   4491: 'Carrier 70 Standard Input Card Fault', class No Acknowledgement, trigger "DB302_HMI_Faults_Carrier70_Faults_0" bit 10
   4492: 'Carrier 70 Standard Output Card Fault', class No Acknowledgement, trigger "DB302_HMI_Faults_Carrier70_Faults_0" bit 11
   4493: 'Carrier 70 Encoder Position Fault', class No Acknowledgement, trigger "DB302_HMI_Faults_Carrier70_Faults_0" bit 12
   4494: 'Carrier 70 Encoder Internal Error', class No Acknowledgement, trigger "DB302_HMI_Faults_Carrier70_Faults_0" bit 13
   4495: 'Carrier 70 Encoder Comm Fault', class No Acknowledgement, trigger "DB302_HMI_Faults_Carrier70_Faults_0" bit 14
   4496: 'Carrier 70 HMI Comm Fault', class No Acknowledgement, trigger "DB302_HMI_Faults_Carrier70_Faults_0" bit 15
   4497: 'Carrier 70 Crash Detection Fault', class No Acknowledgement, trigger "DB302_HMI_Faults_Carrier70_Faults_1" bit 0
   4498: 'Carrier 70 Carrier Number Invalid', class No Acknowledgement, trigger "DB302_HMI_Faults_Carrier70_Faults_1" bit 1
   4499: 'Carrier 70 Drive: PROFINET configuration error', class No Acknowledgement, trigger "DB302_HMI_Faults_Carrier70_Faults_1" bit 2
   4500: 'Carrier 70 Drive: Error internal communications', class No Acknowledgement, trigger "DB302_HMI_Faults_Carrier70_Faults_1" bit 3
   4501: 'Carrier 70 Drive: Motor overtemperature', class No Acknowledgement, trigger "DB302_HMI_Faults_Carrier70_Faults_1" bit 4
   4502: 'Carrier 70 Drive: Motor overcurrent', class No Acknowledgement, trigger "DB302_HMI_Faults_Carrier70_Faults_1" bit 5
   4503: 'Carrier 70 Drive: Infeed or power unit not ready', class No Acknowledgement, trigger "DB302_HMI_Faults_Carrier70_Faults_1" bit 6
   4504: 'Carrier 70 Drive: Short-circuit/ground fault detected', class No Acknowledgement, trigger "DB302_HMI_Faults_Carrier70_Faults_1" bit 7
   4505: 'Carrier 70 Drive: PROFINET Setpoint timeout', class No Acknowledgement, trigger "DB302_HMI_Faults_Carrier70_Faults_1" bit 8
   4506: 'Carrier 70 Power unit: Overcurrent', class No Acknowledgement, trigger "DB302_HMI_Faults_Carrier70_Faults_1" bit 9
   4507: 'Carrier 70 Power unit: DC link voltage overvoltage', class No Acknowledgement, trigger "DB302_HMI_Faults_Carrier70_Faults_1" bit 10
   4508: 'Carrier 70 Power unit: DC link voltage undervoltage', class No Acknowledgement, trigger "DB302_HMI_Faults_Carrier70_Faults_1" bit 11
   4509: 'Carrier 70 Power unit: Line phase failure in main circuit', class No Acknowledgement, trigger "DB302_HMI_Faults_Carrier70_Faults_1" bit 12
   4510: 'Carrier 70 Power unit: Phase failure motor cable', class No Acknowledgement, trigger "DB302_HMI_Faults_Carrier70_Faults_1" bit 13
   4511: 'Carrier 70 Power unit: Ground fault', class No Acknowledgement, trigger "DB302_HMI_Faults_Carrier70_Faults_1" bit 14
   4512: 'Spare_Fault_4512', class No Acknowledgement, trigger "DB302_HMI_Faults_Carrier70_Faults_1" bit 15
   4513: 'Carrier 70 Motion Off Fault', class No Acknowledgement, trigger "DB302_HMI_Faults_Carrier70_Faults_2" bit 0
   4514: 'Carrier 70 Motion On Fault', class No Acknowledgement, trigger "DB302_HMI_Faults_Carrier70_Faults_2" bit 1
   4515: 'Carrier 70 Spacing Fault', class No Acknowledgement, trigger "DB302_HMI_Faults_Carrier70_Faults_2" bit 2
   4516: 'Carrier 70 Duplicate Carrier Number Fault', class No Acknowledgement, trigger "DB302_HMI_Faults_Carrier70_Faults_2" bit 3
   4517: 'Spare_Fault_4517', class No Acknowledgement, trigger "DB302_HMI_Faults_Carrier70_Faults_2" bit 4
   4518: 'Spare_Fault_4518', class No Acknowledgement, trigger "DB302_HMI_Faults_Carrier70_Faults_2" bit 5
   4519: 'Spare_Fault_4519', class No Acknowledgement, trigger "DB302_HMI_Faults_Carrier70_Faults_2" bit 6
   4520: 'Spare_Fault_4520', class No Acknowledgement, trigger "DB302_HMI_Faults_Carrier70_Faults_2" bit 7
   4521: 'Spare_Fault_4521', class No Acknowledgement, trigger "DB302_HMI_Faults_Carrier70_Faults_2" bit 8
   4522: 'Spare_Fault_4522', class No Acknowledgement, trigger "DB302_HMI_Faults_Carrier70_Faults_2" bit 9
   4523: 'Spare_Fault_4523', class No Acknowledgement, trigger "DB302_HMI_Faults_Carrier70_Faults_2" bit 10
   4524: 'Spare_Fault_4524', class No Acknowledgement, trigger "DB302_HMI_Faults_Carrier70_Faults_2" bit 11
   4525: 'Spare_Fault_4525', class No Acknowledgement, trigger "DB302_HMI_Faults_Carrier70_Faults_2" bit 12
   4526: 'Spare_Fault_4526', class No Acknowledgement, trigger "DB302_HMI_Faults_Carrier70_Faults_2" bit 13
   4527: 'Spare_Fault_4527', class No Acknowledgement, trigger "DB302_HMI_Faults_Carrier70_Faults_2" bit 14
   4528: 'Spare_Fault_4528', class No Acknowledgement, trigger "DB302_HMI_Faults_Carrier70_Faults_2" bit 15
   4529: 'Spare_Fault_4529', class No Acknowledgement, trigger "DB302_HMI_Faults_Carrier70_Faults_3" bit 0
   4530: 'Spare_Fault_4530', class No Acknowledgement, trigger "DB302_HMI_Faults_Carrier70_Faults_3" bit 1
   4531: 'Spare_Fault_4531', class No Acknowledgement, trigger "DB302_HMI_Faults_Carrier70_Faults_3" bit 2
   4532: 'Spare_Fault_4532', class No Acknowledgement, trigger "DB302_HMI_Faults_Carrier70_Faults_3" bit 3
   4533: 'Spare_Fault_4533', class No Acknowledgement, trigger "DB302_HMI_Faults_Carrier70_Faults_3" bit 4
   4534: 'Spare_Fault_4534', class No Acknowledgement, trigger "DB302_HMI_Faults_Carrier70_Faults_3" bit 5
   4535: 'Spare_Fault_4535', class No Acknowledgement, trigger "DB302_HMI_Faults_Carrier70_Faults_3" bit 6
   4536: 'Spare_Fault_4536', class No Acknowledgement, trigger "DB302_HMI_Faults_Carrier70_Faults_3" bit 7
   4537: 'Spare_Fault_4537', class No Acknowledgement, trigger "DB302_HMI_Faults_Carrier70_Faults_3" bit 8
   4538: 'Spare_Fault_4538', class No Acknowledgement, trigger "DB302_HMI_Faults_Carrier70_Faults_3" bit 9
   4539: 'Spare_Fault_4539', class No Acknowledgement, trigger "DB302_HMI_Faults_Carrier70_Faults_3" bit 10
   4540: 'Spare_Fault_4540', class No Acknowledgement, trigger "DB302_HMI_Faults_Carrier70_Faults_3" bit 11
   4541: 'Spare_Fault_4541', class No Acknowledgement, trigger "DB302_HMI_Faults_Carrier70_Faults_3" bit 12
   4542: 'Spare_Fault_4542', class No Acknowledgement, trigger "DB302_HMI_Faults_Carrier70_Faults_3" bit 13
   4543: 'Spare_Fault_4543', class No Acknowledgement, trigger "DB302_HMI_Faults_Carrier70_Faults_3" bit 14
   4544: 'Spare_Fault_4544', class No Acknowledgement, trigger "DB302_HMI_Faults_Carrier70_Faults_3" bit 15
   4545: 'Carrier 71 Disconnect Open Power Fault DI11.0', class No Acknowledgement, trigger "DB302_HMI_Faults_Carrier71_Faults_0" bit 0
   4546: 'Carrier 71 Drive Profinet Comm Fault', class No Acknowledgement, trigger "DB302_HMI_Faults_Carrier71_Faults_0" bit 1
   4547: 'Carrier 71 Production Stop Not Reset', class No Acknowledgement, trigger "DB302_HMI_Faults_Carrier71_Faults_0" bit 2
   4548: 'Carrier 71 CB02122 Tripped', class No Acknowledgement, trigger "DB302_HMI_Faults_Carrier71_Faults_0" bit 3
   4549: 'Carrier 71 CB02123 Tripped', class No Acknowledgement, trigger "DB302_HMI_Faults_Carrier71_Faults_0" bit 4
   4550: 'Carrier 71 AUX1 CB Tripped', class No Acknowledgement, trigger "DB302_HMI_Faults_Carrier71_Faults_0" bit 5
   4551: 'Carrier 71 AUX2 CB Tripped', class No Acknowledgement, trigger "DB302_HMI_Faults_Carrier71_Faults_0" bit 6
   4552: 'Carrier 71 PLC Not Communicating', class No Acknowledgement, trigger "DB302_HMI_Faults_Carrier71_Faults_0" bit 7
   4553: 'Carrier 71 Safe Input Card Fault', class No Acknowledgement, trigger "DB302_HMI_Faults_Carrier71_Faults_0" bit 8
   4554: 'Carrier 71 Safe Output Card Fault', class No Acknowledgement, trigger "DB302_HMI_Faults_Carrier71_Faults_0" bit 9
   4555: 'Carrier 71 Standard Input Card Fault', class No Acknowledgement, trigger "DB302_HMI_Faults_Carrier71_Faults_0" bit 10
   4556: 'Carrier 71 Standard Output Card Fault', class No Acknowledgement, trigger "DB302_HMI_Faults_Carrier71_Faults_0" bit 11
   4557: 'Carrier 71 Encoder Position Fault', class No Acknowledgement, trigger "DB302_HMI_Faults_Carrier71_Faults_0" bit 12
   4558: 'Carrier 71 Encoder Internal Error', class No Acknowledgement, trigger "DB302_HMI_Faults_Carrier71_Faults_0" bit 13
   4559: 'Carrier 71 Encoder Comm Fault', class No Acknowledgement, trigger "DB302_HMI_Faults_Carrier71_Faults_0" bit 14
   4560: 'Carrier 71 HMI Comm Fault', class No Acknowledgement, trigger "DB302_HMI_Faults_Carrier71_Faults_0" bit 15
   4561: 'Carrier 71 Crash Detection Fault', class No Acknowledgement, trigger "DB302_HMI_Faults_Carrier71_Faults_1" bit 0
   4562: 'Carrier 71 Carrier Number Invalid', class No Acknowledgement, trigger "DB302_HMI_Faults_Carrier71_Faults_1" bit 1
   4563: 'Carrier 71 Drive: PROFINET configuration error', class No Acknowledgement, trigger "DB302_HMI_Faults_Carrier71_Faults_1" bit 2
   4564: 'Carrier 71 Drive: Error internal communications', class No Acknowledgement, trigger "DB302_HMI_Faults_Carrier71_Faults_1" bit 3
   4565: 'Carrier 71 Drive: Motor overtemperature', class No Acknowledgement, trigger "DB302_HMI_Faults_Carrier71_Faults_1" bit 4
   4566: 'Carrier 71 Drive: Motor overcurrent', class No Acknowledgement, trigger "DB302_HMI_Faults_Carrier71_Faults_1" bit 5
   4567: 'Carrier 71 Drive: Infeed or power unit not ready', class No Acknowledgement, trigger "DB302_HMI_Faults_Carrier71_Faults_1" bit 6
   4568: 'Carrier 71 Drive: Short-circuit/ground fault detected', class No Acknowledgement, trigger "DB302_HMI_Faults_Carrier71_Faults_1" bit 7
   4569: 'Carrier 71 Drive: PROFINET Setpoint timeout', class No Acknowledgement, trigger "DB302_HMI_Faults_Carrier71_Faults_1" bit 8
   4570: 'Carrier 71 Power unit: Overcurrent', class No Acknowledgement, trigger "DB302_HMI_Faults_Carrier71_Faults_1" bit 9
   4571: 'Carrier 71 Power unit: DC link voltage overvoltage', class No Acknowledgement, trigger "DB302_HMI_Faults_Carrier71_Faults_1" bit 10
   4572: 'Carrier 71 Power unit: DC link voltage undervoltage', class No Acknowledgement, trigger "DB302_HMI_Faults_Carrier71_Faults_1" bit 11
   4573: 'Carrier 71 Power unit: Line phase failure in main circuit', class No Acknowledgement, trigger "DB302_HMI_Faults_Carrier71_Faults_1" bit 12
   4574: 'Carrier 71 Power unit: Phase failure motor cable', class No Acknowledgement, trigger "DB302_HMI_Faults_Carrier71_Faults_1" bit 13
   4575: 'Carrier 71 Power unit: Ground fault', class No Acknowledgement, trigger "DB302_HMI_Faults_Carrier71_Faults_1" bit 14
   4576: 'Spare_Fault_4576', class No Acknowledgement, trigger "DB302_HMI_Faults_Carrier71_Faults_1" bit 15
   4577: 'Carrier 71 Motion Off Fault', class No Acknowledgement, trigger "DB302_HMI_Faults_Carrier71_Faults_2" bit 0
   4578: 'Carrier 71 Motion On Fault', class No Acknowledgement, trigger "DB302_HMI_Faults_Carrier71_Faults_2" bit 1
   4579: 'Carrier 71 Spacing Fault', class No Acknowledgement, trigger "DB302_HMI_Faults_Carrier71_Faults_2" bit 2
   4580: 'Carrier 71 Duplicate Carrier Number Fault', class No Acknowledgement, trigger "DB302_HMI_Faults_Carrier71_Faults_2" bit 3
   4581: 'Spare_Fault_4581', class No Acknowledgement, trigger "DB302_HMI_Faults_Carrier71_Faults_2" bit 4
   4582: 'Spare_Fault_4582', class No Acknowledgement, trigger "DB302_HMI_Faults_Carrier71_Faults_2" bit 5
   4583: 'Spare_Fault_4583', class No Acknowledgement, trigger "DB302_HMI_Faults_Carrier71_Faults_2" bit 6
   4584: 'Spare_Fault_4584', class No Acknowledgement, trigger "DB302_HMI_Faults_Carrier71_Faults_2" bit 7
   4585: 'Spare_Fault_4585', class No Acknowledgement, trigger "DB302_HMI_Faults_Carrier71_Faults_2" bit 8
   4586: 'Spare_Fault_4586', class No Acknowledgement, trigger "DB302_HMI_Faults_Carrier71_Faults_2" bit 9
   4587: 'Spare_Fault_4587', class No Acknowledgement, trigger "DB302_HMI_Faults_Carrier71_Faults_2" bit 10
   4588: 'Spare_Fault_4588', class No Acknowledgement, trigger "DB302_HMI_Faults_Carrier71_Faults_2" bit 11
   4589: 'Spare_Fault_4589', class No Acknowledgement, trigger "DB302_HMI_Faults_Carrier71_Faults_2" bit 12
   4590: 'Spare_Fault_4590', class No Acknowledgement, trigger "DB302_HMI_Faults_Carrier71_Faults_2" bit 13
   4591: 'Spare_Fault_4591', class No Acknowledgement, trigger "DB302_HMI_Faults_Carrier71_Faults_2" bit 14
   4592: 'Spare_Fault_4592', class No Acknowledgement, trigger "DB302_HMI_Faults_Carrier71_Faults_2" bit 15
   4593: 'Spare_Fault_4593', class No Acknowledgement, trigger "DB302_HMI_Faults_Carrier71_Faults_3" bit 0
   4594: 'Spare_Fault_4594', class No Acknowledgement, trigger "DB302_HMI_Faults_Carrier71_Faults_3" bit 1
   4595: 'Spare_Fault_4595', class No Acknowledgement, trigger "DB302_HMI_Faults_Carrier71_Faults_3" bit 2
   4596: 'Spare_Fault_4596', class No Acknowledgement, trigger "DB302_HMI_Faults_Carrier71_Faults_3" bit 3
   4597: 'Spare_Fault_4597', class No Acknowledgement, trigger "DB302_HMI_Faults_Carrier71_Faults_3" bit 4
   4598: 'Spare_Fault_4598', class No Acknowledgement, trigger "DB302_HMI_Faults_Carrier71_Faults_3" bit 5
   4599: 'Spare_Fault_4599', class No Acknowledgement, trigger "DB302_HMI_Faults_Carrier71_Faults_3" bit 6
   4600: 'Spare_Fault_4600', class No Acknowledgement, trigger "DB302_HMI_Faults_Carrier71_Faults_3" bit 7
   4601: 'Spare_Fault_4601', class No Acknowledgement, trigger "DB302_HMI_Faults_Carrier71_Faults_3" bit 8
   4602: 'Spare_Fault_4602', class No Acknowledgement, trigger "DB302_HMI_Faults_Carrier71_Faults_3" bit 9
   4603: 'Spare_Fault_4603', class No Acknowledgement, trigger "DB302_HMI_Faults_Carrier71_Faults_3" bit 10
   4604: 'Spare_Fault_4604', class No Acknowledgement, trigger "DB302_HMI_Faults_Carrier71_Faults_3" bit 11
   4605: 'Spare_Fault_4605', class No Acknowledgement, trigger "DB302_HMI_Faults_Carrier71_Faults_3" bit 12
   4606: 'Spare_Fault_4606', class No Acknowledgement, trigger "DB302_HMI_Faults_Carrier71_Faults_3" bit 13
   4607: 'Spare_Fault_4607', class No Acknowledgement, trigger "DB302_HMI_Faults_Carrier71_Faults_3" bit 14
   4608: 'Spare_Fault_4608', class No Acknowledgement, trigger "DB302_HMI_Faults_Carrier71_Faults_3" bit 15
   4609: 'Carrier 72 Disconnect Open Power Fault DI11.0', class No Acknowledgement, trigger "DB302_HMI_Faults_Carrier72_Faults_0" bit 0
   4610: 'Carrier 72 Drive Profinet Comm Fault', class No Acknowledgement, trigger "DB302_HMI_Faults_Carrier72_Faults_0" bit 1
   4611: 'Carrier 72 Production Stop Not Reset', class No Acknowledgement, trigger "DB302_HMI_Faults_Carrier72_Faults_0" bit 2
   4612: 'Carrier 72 CB02122 Tripped', class No Acknowledgement, trigger "DB302_HMI_Faults_Carrier72_Faults_0" bit 3
   4613: 'Carrier 72 CB02123 Tripped', class No Acknowledgement, trigger "DB302_HMI_Faults_Carrier72_Faults_0" bit 4
   4614: 'Carrier 72 AUX1 CB Tripped', class No Acknowledgement, trigger "DB302_HMI_Faults_Carrier72_Faults_0" bit 5
   4615: 'Carrier 72 AUX2 CB Tripped', class No Acknowledgement, trigger "DB302_HMI_Faults_Carrier72_Faults_0" bit 6
   4616: 'Carrier 72 PLC Not Communicating', class No Acknowledgement, trigger "DB302_HMI_Faults_Carrier72_Faults_0" bit 7
   4617: 'Carrier 72 Safe Input Card Fault', class No Acknowledgement, trigger "DB302_HMI_Faults_Carrier72_Faults_0" bit 8
   4618: 'Carrier 72 Safe Output Card Fault', class No Acknowledgement, trigger "DB302_HMI_Faults_Carrier72_Faults_0" bit 9
   4619: 'Carrier 72 Standard Input Card Fault', class No Acknowledgement, trigger "DB302_HMI_Faults_Carrier72_Faults_0" bit 10
   4620: 'Carrier 72 Standard Output Card Fault', class No Acknowledgement, trigger "DB302_HMI_Faults_Carrier72_Faults_0" bit 11
   4621: 'Carrier 72 Encoder Position Fault', class No Acknowledgement, trigger "DB302_HMI_Faults_Carrier72_Faults_0" bit 12
   4622: 'Carrier 72 Encoder Internal Error', class No Acknowledgement, trigger "DB302_HMI_Faults_Carrier72_Faults_0" bit 13
   4623: 'Carrier 72 Encoder Comm Fault', class No Acknowledgement, trigger "DB302_HMI_Faults_Carrier72_Faults_0" bit 14
   4624: 'Carrier 72 HMI Comm Fault', class No Acknowledgement, trigger "DB302_HMI_Faults_Carrier72_Faults_0" bit 15
   4625: 'Carrier 72 Crash Detection Fault', class No Acknowledgement, trigger "DB302_HMI_Faults_Carrier72_Faults_1" bit 0
   4626: 'Carrier 72 Carrier Number Invalid', class No Acknowledgement, trigger "DB302_HMI_Faults_Carrier72_Faults_1" bit 1
   4627: 'Carrier 72 Drive: PROFINET configuration error', class No Acknowledgement, trigger "DB302_HMI_Faults_Carrier72_Faults_1" bit 2
   4628: 'Carrier 72 Drive: Error internal communications', class No Acknowledgement, trigger "DB302_HMI_Faults_Carrier72_Faults_1" bit 3
   4629: 'Carrier 72 Drive: Motor overtemperature', class No Acknowledgement, trigger "DB302_HMI_Faults_Carrier72_Faults_1" bit 4
   4630: 'Carrier 72 Drive: Motor overcurrent', class No Acknowledgement, trigger "DB302_HMI_Faults_Carrier72_Faults_1" bit 5
   4631: 'Carrier 72 Drive: Infeed or power unit not ready', class No Acknowledgement, trigger "DB302_HMI_Faults_Carrier72_Faults_1" bit 6
   4632: 'Carrier 72 Drive: Short-circuit/ground fault detected', class No Acknowledgement, trigger "DB302_HMI_Faults_Carrier72_Faults_1" bit 7
   4633: 'Carrier 72 Drive: PROFINET Setpoint timeout', class No Acknowledgement, trigger "DB302_HMI_Faults_Carrier72_Faults_1" bit 8
   4634: 'Carrier 72 Power unit: Overcurrent', class No Acknowledgement, trigger "DB302_HMI_Faults_Carrier72_Faults_1" bit 9
   4635: 'Carrier 72 Power unit: DC link voltage overvoltage', class No Acknowledgement, trigger "DB302_HMI_Faults_Carrier72_Faults_1" bit 10
   4636: 'Carrier 72 Power unit: DC link voltage undervoltage', class No Acknowledgement, trigger "DB302_HMI_Faults_Carrier72_Faults_1" bit 11
   4637: 'Carrier 72 Power unit: Line phase failure in main circuit', class No Acknowledgement, trigger "DB302_HMI_Faults_Carrier72_Faults_1" bit 12
   4638: 'Carrier 72 Power unit: Phase failure motor cable', class No Acknowledgement, trigger "DB302_HMI_Faults_Carrier72_Faults_1" bit 13
   4639: 'Carrier 72 Power unit: Ground fault', class No Acknowledgement, trigger "DB302_HMI_Faults_Carrier72_Faults_1" bit 14
   4640: 'Spare_Fault_4640', class No Acknowledgement, trigger "DB302_HMI_Faults_Carrier72_Faults_1" bit 15
   4641: 'Carrier 72 Motion Off Fault', class No Acknowledgement, trigger "DB302_HMI_Faults_Carrier72_Faults_2" bit 0
   4642: 'Carrier 72 Motion On Fault', class No Acknowledgement, trigger "DB302_HMI_Faults_Carrier72_Faults_2" bit 1
   4643: 'Carrier 72 Spacing Fault', class No Acknowledgement, trigger "DB302_HMI_Faults_Carrier72_Faults_2" bit 2
   4644: 'Carrier 72 Duplicate Carrier Number Fault', class No Acknowledgement, trigger "DB302_HMI_Faults_Carrier72_Faults_2" bit 3
   4645: 'Spare_Fault_4645', class No Acknowledgement, trigger "DB302_HMI_Faults_Carrier72_Faults_2" bit 4
   4646: 'Spare_Fault_4646', class No Acknowledgement, trigger "DB302_HMI_Faults_Carrier72_Faults_2" bit 5
   4647: 'Spare_Fault_4647', class No Acknowledgement, trigger "DB302_HMI_Faults_Carrier72_Faults_2" bit 6
   4648: 'Spare_Fault_4648', class No Acknowledgement, trigger "DB302_HMI_Faults_Carrier72_Faults_2" bit 7
   4649: 'Spare_Fault_4649', class No Acknowledgement, trigger "DB302_HMI_Faults_Carrier72_Faults_2" bit 8
   4650: 'Spare_Fault_4650', class No Acknowledgement, trigger "DB302_HMI_Faults_Carrier72_Faults_2" bit 9
   4651: 'Spare_Fault_4651', class No Acknowledgement, trigger "DB302_HMI_Faults_Carrier72_Faults_2" bit 10
   4652: 'Spare_Fault_4652', class No Acknowledgement, trigger "DB302_HMI_Faults_Carrier72_Faults_2" bit 11
   4653: 'Spare_Fault_4653', class No Acknowledgement, trigger "DB302_HMI_Faults_Carrier72_Faults_2" bit 12
   4654: 'Spare_Fault_4654', class No Acknowledgement, trigger "DB302_HMI_Faults_Carrier72_Faults_2" bit 13
   4655: 'Spare_Fault_4655', class No Acknowledgement, trigger "DB302_HMI_Faults_Carrier72_Faults_2" bit 14
   4656: 'Spare_Fault_4656', class No Acknowledgement, trigger "DB302_HMI_Faults_Carrier72_Faults_2" bit 15
   4657: 'Spare_Fault_4657', class No Acknowledgement, trigger "DB302_HMI_Faults_Carrier72_Faults_3" bit 0
   4658: 'Spare_Fault_4658', class No Acknowledgement, trigger "DB302_HMI_Faults_Carrier72_Faults_3" bit 1
   4659: 'Spare_Fault_4659', class No Acknowledgement, trigger "DB302_HMI_Faults_Carrier72_Faults_3" bit 2
   4660: 'Spare_Fault_4660', class No Acknowledgement, trigger "DB302_HMI_Faults_Carrier72_Faults_3" bit 3
   4661: 'Spare_Fault_4661', class No Acknowledgement, trigger "DB302_HMI_Faults_Carrier72_Faults_3" bit 4
   4662: 'Spare_Fault_4662', class No Acknowledgement, trigger "DB302_HMI_Faults_Carrier72_Faults_3" bit 5
   4663: 'Spare_Fault_4663', class No Acknowledgement, trigger "DB302_HMI_Faults_Carrier72_Faults_3" bit 6
   4664: 'Spare_Fault_4664', class No Acknowledgement, trigger "DB302_HMI_Faults_Carrier72_Faults_3" bit 7
   4665: 'Spare_Fault_4665', class No Acknowledgement, trigger "DB302_HMI_Faults_Carrier72_Faults_3" bit 8
   4666: 'Spare_Fault_4666', class No Acknowledgement, trigger "DB302_HMI_Faults_Carrier72_Faults_3" bit 9
   4667: 'Spare_Fault_4667', class No Acknowledgement, trigger "DB302_HMI_Faults_Carrier72_Faults_3" bit 10
   4668: 'Spare_Fault_4668', class No Acknowledgement, trigger "DB302_HMI_Faults_Carrier72_Faults_3" bit 11
   4669: 'Spare_Fault_4669', class No Acknowledgement, trigger "DB302_HMI_Faults_Carrier72_Faults_3" bit 12
   4670: 'Spare_Fault_4670', class No Acknowledgement, trigger "DB302_HMI_Faults_Carrier72_Faults_3" bit 13
   4671: 'Spare_Fault_4671', class No Acknowledgement, trigger "DB302_HMI_Faults_Carrier72_Faults_3" bit 14
   4672: 'Spare_Fault_4672', class No Acknowledgement, trigger "DB302_HMI_Faults_Carrier72_Faults_3" bit 15
   4673: 'Carrier 73 Disconnect Open Power Fault DI11.0', class No Acknowledgement, trigger "DB302_HMI_Faults_Carrier73_Faults_0" bit 0
   4674: 'Carrier 73 Drive Profinet Comm Fault', class No Acknowledgement, trigger "DB302_HMI_Faults_Carrier73_Faults_0" bit 1
   4675: 'Carrier 73 Production Stop Not Reset', class No Acknowledgement, trigger "DB302_HMI_Faults_Carrier73_Faults_0" bit 2
   4676: 'Carrier 73 CB02122 Tripped', class No Acknowledgement, trigger "DB302_HMI_Faults_Carrier73_Faults_0" bit 3
   4677: 'Carrier 73 CB02123 Tripped', class No Acknowledgement, trigger "DB302_HMI_Faults_Carrier73_Faults_0" bit 4
   4678: 'Carrier 73 AUX1 CB Tripped', class No Acknowledgement, trigger "DB302_HMI_Faults_Carrier73_Faults_0" bit 5
   4679: 'Carrier 73 AUX2 CB Tripped', class No Acknowledgement, trigger "DB302_HMI_Faults_Carrier73_Faults_0" bit 6
   4680: 'Carrier 73 PLC Not Communicating', class No Acknowledgement, trigger "DB302_HMI_Faults_Carrier73_Faults_0" bit 7
   4681: 'Carrier 73 Safe Input Card Fault', class No Acknowledgement, trigger "DB302_HMI_Faults_Carrier73_Faults_0" bit 8
   4682: 'Carrier 73 Safe Output Card Fault', class No Acknowledgement, trigger "DB302_HMI_Faults_Carrier73_Faults_0" bit 9
   4683: 'Carrier 73 Standard Input Card Fault', class No Acknowledgement, trigger "DB302_HMI_Faults_Carrier73_Faults_0" bit 10
   4684: 'Carrier 73 Standard Output Card Fault', class No Acknowledgement, trigger "DB302_HMI_Faults_Carrier73_Faults_0" bit 11
   4685: 'Carrier 73 Encoder Position Fault', class No Acknowledgement, trigger "DB302_HMI_Faults_Carrier73_Faults_0" bit 12
   4686: 'Carrier 73 Encoder Internal Error', class No Acknowledgement, trigger "DB302_HMI_Faults_Carrier73_Faults_0" bit 13
   4687: 'Carrier 73 Encoder Comm Fault', class No Acknowledgement, trigger "DB302_HMI_Faults_Carrier73_Faults_0" bit 14
   4688: 'Carrier 73 HMI Comm Fault', class No Acknowledgement, trigger "DB302_HMI_Faults_Carrier73_Faults_0" bit 15
   4689: 'Carrier 73 Crash Detection Fault', class No Acknowledgement, trigger "DB302_HMI_Faults_Carrier73_Faults_1" bit 0
   4690: 'Carrier 73 Carrier Number Invalid', class No Acknowledgement, trigger "DB302_HMI_Faults_Carrier73_Faults_1" bit 1
   4691: 'Carrier 73 Drive: PROFINET configuration error', class No Acknowledgement, trigger "DB302_HMI_Faults_Carrier73_Faults_1" bit 2
   4692: 'Carrier 73 Drive: Error internal communications', class No Acknowledgement, trigger "DB302_HMI_Faults_Carrier73_Faults_1" bit 3
   4693: 'Carrier 73 Drive: Motor overtemperature', class No Acknowledgement, trigger "DB302_HMI_Faults_Carrier73_Faults_1" bit 4
   4694: 'Carrier 73 Drive: Motor overcurrent', class No Acknowledgement, trigger "DB302_HMI_Faults_Carrier73_Faults_1" bit 5
   4695: 'Carrier 73 Drive: Infeed or power unit not ready', class No Acknowledgement, trigger "DB302_HMI_Faults_Carrier73_Faults_1" bit 6
   4696: 'Carrier 73 Drive: Short-circuit/ground fault detected', class No Acknowledgement, trigger "DB302_HMI_Faults_Carrier73_Faults_1" bit 7
   4697: 'Carrier 73 Drive: PROFINET Setpoint timeout', class No Acknowledgement, trigger "DB302_HMI_Faults_Carrier73_Faults_1" bit 8
   4698: 'Carrier 73 Power unit: Overcurrent', class No Acknowledgement, trigger "DB302_HMI_Faults_Carrier73_Faults_1" bit 9
   4699: 'Carrier 73 Power unit: DC link voltage overvoltage', class No Acknowledgement, trigger "DB302_HMI_Faults_Carrier73_Faults_1" bit 10
   4700: 'Carrier 73 Power unit: DC link voltage undervoltage', class No Acknowledgement, trigger "DB302_HMI_Faults_Carrier73_Faults_1" bit 11
   4701: 'Carrier 73 Power unit: Line phase failure in main circuit', class No Acknowledgement, trigger "DB302_HMI_Faults_Carrier73_Faults_1" bit 12
   4702: 'Carrier 73 Power unit: Phase failure motor cable', class No Acknowledgement, trigger "DB302_HMI_Faults_Carrier73_Faults_1" bit 13
   4703: 'Carrier 73 Power unit: Ground fault', class No Acknowledgement, trigger "DB302_HMI_Faults_Carrier73_Faults_1" bit 14
   4704: 'Spare_Fault_4704', class No Acknowledgement, trigger "DB302_HMI_Faults_Carrier73_Faults_1" bit 15
   4705: 'Carrier 73 Motion Off Fault', class No Acknowledgement, trigger "DB302_HMI_Faults_Carrier73_Faults_2" bit 0
   4706: 'Carrier 73 Motion On Fault', class No Acknowledgement, trigger "DB302_HMI_Faults_Carrier73_Faults_2" bit 1
   4707: 'Carrier 73 Spacing Fault', class No Acknowledgement, trigger "DB302_HMI_Faults_Carrier73_Faults_2" bit 2
   4708: 'Carrier 73 Duplicate Carrier Number Fault', class No Acknowledgement, trigger "DB302_HMI_Faults_Carrier73_Faults_2" bit 3
   4709: 'Spare_Fault_4709', class No Acknowledgement, trigger "DB302_HMI_Faults_Carrier73_Faults_2" bit 4
   4710: 'Spare_Fault_4710', class No Acknowledgement, trigger "DB302_HMI_Faults_Carrier73_Faults_2" bit 5
   4711: 'Spare_Fault_4711', class No Acknowledgement, trigger "DB302_HMI_Faults_Carrier73_Faults_2" bit 6
   4712: 'Spare_Fault_4712', class No Acknowledgement, trigger "DB302_HMI_Faults_Carrier73_Faults_2" bit 7
   4713: 'Spare_Fault_4713', class No Acknowledgement, trigger "DB302_HMI_Faults_Carrier73_Faults_2" bit 8
   4714: 'Spare_Fault_4714', class No Acknowledgement, trigger "DB302_HMI_Faults_Carrier73_Faults_2" bit 9
   4715: 'Spare_Fault_4715', class No Acknowledgement, trigger "DB302_HMI_Faults_Carrier73_Faults_2" bit 10
   4716: 'Spare_Fault_4716', class No Acknowledgement, trigger "DB302_HMI_Faults_Carrier73_Faults_2" bit 11
   4717: 'Spare_Fault_4717', class No Acknowledgement, trigger "DB302_HMI_Faults_Carrier73_Faults_2" bit 12
   4718: 'Spare_Fault_4718', class No Acknowledgement, trigger "DB302_HMI_Faults_Carrier73_Faults_2" bit 13
   4719: 'Spare_Fault_4719', class No Acknowledgement, trigger "DB302_HMI_Faults_Carrier73_Faults_2" bit 14
   4720: 'Spare_Fault_4720', class No Acknowledgement, trigger "DB302_HMI_Faults_Carrier73_Faults_2" bit 15
   4721: 'Spare_Fault_4721', class No Acknowledgement, trigger "DB302_HMI_Faults_Carrier73_Faults_3" bit 0
   4722: 'Spare_Fault_4722', class No Acknowledgement, trigger "DB302_HMI_Faults_Carrier73_Faults_3" bit 1
   4723: 'Spare_Fault_4723', class No Acknowledgement, trigger "DB302_HMI_Faults_Carrier73_Faults_3" bit 2
   4724: 'Spare_Fault_4724', class No Acknowledgement, trigger "DB302_HMI_Faults_Carrier73_Faults_3" bit 3
   4725: 'Spare_Fault_4725', class No Acknowledgement, trigger "DB302_HMI_Faults_Carrier73_Faults_3" bit 4
   4726: 'Spare_Fault_4726', class No Acknowledgement, trigger "DB302_HMI_Faults_Carrier73_Faults_3" bit 5
   4727: 'Spare_Fault_4727', class No Acknowledgement, trigger "DB302_HMI_Faults_Carrier73_Faults_3" bit 6
   4728: 'Spare_Fault_4728', class No Acknowledgement, trigger "DB302_HMI_Faults_Carrier73_Faults_3" bit 7
   4729: 'Spare_Fault_4729', class No Acknowledgement, trigger "DB302_HMI_Faults_Carrier73_Faults_3" bit 8
   4730: 'Spare_Fault_4730', class No Acknowledgement, trigger "DB302_HMI_Faults_Carrier73_Faults_3" bit 9
   4731: 'Spare_Fault_4731', class No Acknowledgement, trigger "DB302_HMI_Faults_Carrier73_Faults_3" bit 10
   4732: 'Spare_Fault_4732', class No Acknowledgement, trigger "DB302_HMI_Faults_Carrier73_Faults_3" bit 11
   4733: 'Spare_Fault_4733', class No Acknowledgement, trigger "DB302_HMI_Faults_Carrier73_Faults_3" bit 12
   4734: 'Spare_Fault_4734', class No Acknowledgement, trigger "DB302_HMI_Faults_Carrier73_Faults_3" bit 13
   4735: 'Spare_Fault_4735', class No Acknowledgement, trigger "DB302_HMI_Faults_Carrier73_Faults_3" bit 14
   4736: 'Spare_Fault_4736', class No Acknowledgement, trigger "DB302_HMI_Faults_Carrier73_Faults_3" bit 15
   4737: 'Carrier 74 Disconnect Open Power Fault DI11.0', class No Acknowledgement, trigger "DB302_HMI_Faults_Carrier74_Faults_0" bit 0
   4738: 'Carrier 74 Drive Profinet Comm Fault', class No Acknowledgement, trigger "DB302_HMI_Faults_Carrier74_Faults_0" bit 1
   4739: 'Carrier 74 Production Stop Not Reset', class No Acknowledgement, trigger "DB302_HMI_Faults_Carrier74_Faults_0" bit 2
   4740: 'Carrier 74 CB02122 Tripped', class No Acknowledgement, trigger "DB302_HMI_Faults_Carrier74_Faults_0" bit 3
   4741: 'Carrier 74 CB02123 Tripped', class No Acknowledgement, trigger "DB302_HMI_Faults_Carrier74_Faults_0" bit 4
   4742: 'Carrier 74 AUX1 CB Tripped', class No Acknowledgement, trigger "DB302_HMI_Faults_Carrier74_Faults_0" bit 5
   4743: 'Carrier 74 AUX2 CB Tripped', class No Acknowledgement, trigger "DB302_HMI_Faults_Carrier74_Faults_0" bit 6
   4744: 'Carrier 74 PLC Not Communicating', class No Acknowledgement, trigger "DB302_HMI_Faults_Carrier74_Faults_0" bit 7
   4745: 'Carrier 74 Safe Input Card Fault', class No Acknowledgement, trigger "DB302_HMI_Faults_Carrier74_Faults_0" bit 8
   4746: 'Carrier 74 Safe Output Card Fault', class No Acknowledgement, trigger "DB302_HMI_Faults_Carrier74_Faults_0" bit 9
   4747: 'Carrier 74 Standard Input Card Fault', class No Acknowledgement, trigger "DB302_HMI_Faults_Carrier74_Faults_0" bit 10
   4748: 'Carrier 74 Standard Output Card Fault', class No Acknowledgement, trigger "DB302_HMI_Faults_Carrier74_Faults_0" bit 11
   4749: 'Carrier 74 Encoder Position Fault', class No Acknowledgement, trigger "DB302_HMI_Faults_Carrier74_Faults_0" bit 12
   4750: 'Carrier 74 Encoder Internal Error', class No Acknowledgement, trigger "DB302_HMI_Faults_Carrier74_Faults_0" bit 13
   4751: 'Carrier 74 Encoder Comm Fault', class No Acknowledgement, trigger "DB302_HMI_Faults_Carrier74_Faults_0" bit 14
   4752: 'Carrier 74 HMI Comm Fault', class No Acknowledgement, trigger "DB302_HMI_Faults_Carrier74_Faults_0" bit 15
   4753: 'Carrier 74 Crash Detection Fault', class No Acknowledgement, trigger "DB302_HMI_Faults_Carrier74_Faults_1" bit 0
   4754: 'Carrier 74 Carrier Number Invalid', class No Acknowledgement, trigger "DB302_HMI_Faults_Carrier74_Faults_1" bit 1
   4755: 'Carrier 74 Drive: PROFINET configuration error', class No Acknowledgement, trigger "DB302_HMI_Faults_Carrier74_Faults_1" bit 2
   4756: 'Carrier 74 Drive: Error internal communications', class No Acknowledgement, trigger "DB302_HMI_Faults_Carrier74_Faults_1" bit 3
   4757: 'Carrier 74 Drive: Motor overtemperature', class No Acknowledgement, trigger "DB302_HMI_Faults_Carrier74_Faults_1" bit 4
   4758: 'Carrier 74 Drive: Motor overcurrent', class No Acknowledgement, trigger "DB302_HMI_Faults_Carrier74_Faults_1" bit 5
   4759: 'Carrier 74 Drive: Infeed or power unit not ready', class No Acknowledgement, trigger "DB302_HMI_Faults_Carrier74_Faults_1" bit 6
   4760: 'Carrier 74 Drive: Short-circuit/ground fault detected', class No Acknowledgement, trigger "DB302_HMI_Faults_Carrier74_Faults_1" bit 7
   4761: 'Carrier 74 Drive: PROFINET Setpoint timeout', class No Acknowledgement, trigger "DB302_HMI_Faults_Carrier74_Faults_1" bit 8
   4762: 'Carrier 74 Power unit: Overcurrent', class No Acknowledgement, trigger "DB302_HMI_Faults_Carrier74_Faults_1" bit 9
   4763: 'Carrier 74 Power unit: DC link voltage overvoltage', class No Acknowledgement, trigger "DB302_HMI_Faults_Carrier74_Faults_1" bit 10
   4764: 'Carrier 74 Power unit: DC link voltage undervoltage', class No Acknowledgement, trigger "DB302_HMI_Faults_Carrier74_Faults_1" bit 11
   4765: 'Carrier 74 Power unit: Line phase failure in main circuit', class No Acknowledgement, trigger "DB302_HMI_Faults_Carrier74_Faults_1" bit 12
   4766: 'Carrier 74 Power unit: Phase failure motor cable', class No Acknowledgement, trigger "DB302_HMI_Faults_Carrier74_Faults_1" bit 13
   4767: 'Carrier 74 Power unit: Ground fault', class No Acknowledgement, trigger "DB302_HMI_Faults_Carrier74_Faults_1" bit 14
   4768: 'Spare_Fault_4768', class No Acknowledgement, trigger "DB302_HMI_Faults_Carrier74_Faults_1" bit 15
   4769: 'Carrier 74 Motion Off Fault', class No Acknowledgement, trigger "DB302_HMI_Faults_Carrier74_Faults_2" bit 0
   4770: 'Carrier 74 Motion On Fault', class No Acknowledgement, trigger "DB302_HMI_Faults_Carrier74_Faults_2" bit 1
   4771: 'Carrier 74 Spacing Fault', class No Acknowledgement, trigger "DB302_HMI_Faults_Carrier74_Faults_2" bit 2
   4772: 'Carrier 74 Duplicate Carrier Number Fault', class No Acknowledgement, trigger "DB302_HMI_Faults_Carrier74_Faults_2" bit 3
   4773: 'Spare_Fault_4773', class No Acknowledgement, trigger "DB302_HMI_Faults_Carrier74_Faults_2" bit 4
   4774: 'Spare_Fault_4774', class No Acknowledgement, trigger "DB302_HMI_Faults_Carrier74_Faults_2" bit 5
   4775: 'Spare_Fault_4775', class No Acknowledgement, trigger "DB302_HMI_Faults_Carrier74_Faults_2" bit 6
   4776: 'Spare_Fault_4776', class No Acknowledgement, trigger "DB302_HMI_Faults_Carrier74_Faults_2" bit 7
   4777: 'Spare_Fault_4777', class No Acknowledgement, trigger "DB302_HMI_Faults_Carrier74_Faults_2" bit 8
   4778: 'Spare_Fault_4778', class No Acknowledgement, trigger "DB302_HMI_Faults_Carrier74_Faults_2" bit 9
   4779: 'Spare_Fault_4779', class No Acknowledgement, trigger "DB302_HMI_Faults_Carrier74_Faults_2" bit 10
   4780: 'Spare_Fault_4780', class No Acknowledgement, trigger "DB302_HMI_Faults_Carrier74_Faults_2" bit 11
   4781: 'Spare_Fault_4781', class No Acknowledgement, trigger "DB302_HMI_Faults_Carrier74_Faults_2" bit 12
   4782: 'Spare_Fault_4782', class No Acknowledgement, trigger "DB302_HMI_Faults_Carrier74_Faults_2" bit 13
   4783: 'Spare_Fault_4783', class No Acknowledgement, trigger "DB302_HMI_Faults_Carrier74_Faults_2" bit 14
   4784: 'Spare_Fault_4784', class No Acknowledgement, trigger "DB302_HMI_Faults_Carrier74_Faults_2" bit 15
   4785: 'Spare_Fault_4785', class No Acknowledgement, trigger "DB302_HMI_Faults_Carrier74_Faults_3" bit 0
   4786: 'Spare_Fault_4786', class No Acknowledgement, trigger "DB302_HMI_Faults_Carrier74_Faults_3" bit 1
   4787: 'Spare_Fault_4787', class No Acknowledgement, trigger "DB302_HMI_Faults_Carrier74_Faults_3" bit 2
   4788: 'Spare_Fault_4788', class No Acknowledgement, trigger "DB302_HMI_Faults_Carrier74_Faults_3" bit 3
   4789: 'Spare_Fault_4789', class No Acknowledgement, trigger "DB302_HMI_Faults_Carrier74_Faults_3" bit 4
   4790: 'Spare_Fault_4790', class No Acknowledgement, trigger "DB302_HMI_Faults_Carrier74_Faults_3" bit 5
   4791: 'Spare_Fault_4791', class No Acknowledgement, trigger "DB302_HMI_Faults_Carrier74_Faults_3" bit 6
   4792: 'Spare_Fault_4792', class No Acknowledgement, trigger "DB302_HMI_Faults_Carrier74_Faults_3" bit 7
   4793: 'Spare_Fault_4793', class No Acknowledgement, trigger "DB302_HMI_Faults_Carrier74_Faults_3" bit 8
   4794: 'Spare_Fault_4794', class No Acknowledgement, trigger "DB302_HMI_Faults_Carrier74_Faults_3" bit 9
   4795: 'Spare_Fault_4795', class No Acknowledgement, trigger "DB302_HMI_Faults_Carrier74_Faults_3" bit 10
   4796: 'Spare_Fault_4796', class No Acknowledgement, trigger "DB302_HMI_Faults_Carrier74_Faults_3" bit 11
   4797: 'Spare_Fault_4797', class No Acknowledgement, trigger "DB302_HMI_Faults_Carrier74_Faults_3" bit 12
   4798: 'Spare_Fault_4798', class No Acknowledgement, trigger "DB302_HMI_Faults_Carrier74_Faults_3" bit 13
   4799: 'Spare_Fault_4799', class No Acknowledgement, trigger "DB302_HMI_Faults_Carrier74_Faults_3" bit 14
   4800: 'Spare_Fault_4800', class No Acknowledgement, trigger "DB302_HMI_Faults_Carrier74_Faults_3" bit 15
   4801: 'Carrier 75 Disconnect Open Power Fault DI11.0', class No Acknowledgement, trigger "DB302_HMI_Faults_Carrier75_Faults_0" bit 0
   4802: 'Carrier 75 Drive Profinet Comm Fault', class No Acknowledgement, trigger "DB302_HMI_Faults_Carrier75_Faults_0" bit 1
   4803: 'Carrier 75 Production Stop Not Reset', class No Acknowledgement, trigger "DB302_HMI_Faults_Carrier75_Faults_0" bit 2
   4804: 'Carrier 75 CB02122 Tripped', class No Acknowledgement, trigger "DB302_HMI_Faults_Carrier75_Faults_0" bit 3
   4805: 'Carrier 75 CB02123 Tripped', class No Acknowledgement, trigger "DB302_HMI_Faults_Carrier75_Faults_0" bit 4
   4806: 'Carrier 75 AUX1 CB Tripped', class No Acknowledgement, trigger "DB302_HMI_Faults_Carrier75_Faults_0" bit 5
   4807: 'Carrier 75 AUX2 CB Tripped', class No Acknowledgement, trigger "DB302_HMI_Faults_Carrier75_Faults_0" bit 6
   4808: 'Carrier 75 PLC Not Communicating', class No Acknowledgement, trigger "DB302_HMI_Faults_Carrier75_Faults_0" bit 7
   4809: 'Carrier 75 Safe Input Card Fault', class No Acknowledgement, trigger "DB302_HMI_Faults_Carrier75_Faults_0" bit 8
   4810: 'Carrier 75 Safe Output Card Fault', class No Acknowledgement, trigger "DB302_HMI_Faults_Carrier75_Faults_0" bit 9
   4811: 'Carrier 75 Standard Input Card Fault', class No Acknowledgement, trigger "DB302_HMI_Faults_Carrier75_Faults_0" bit 10
   4812: 'Carrier 75 Standard Output Card Fault', class No Acknowledgement, trigger "DB302_HMI_Faults_Carrier75_Faults_0" bit 11
   4813: 'Carrier 75 Encoder Position Fault', class No Acknowledgement, trigger "DB302_HMI_Faults_Carrier75_Faults_0" bit 12
   4814: 'Carrier 75 Encoder Internal Error', class No Acknowledgement, trigger "DB302_HMI_Faults_Carrier75_Faults_0" bit 13
   4815: 'Carrier 75 Encoder Comm Fault', class No Acknowledgement, trigger "DB302_HMI_Faults_Carrier75_Faults_0" bit 14
   4816: 'Carrier 75 HMI Comm Fault', class No Acknowledgement, trigger "DB302_HMI_Faults_Carrier75_Faults_0" bit 15
   4817: 'Carrier 75 Crash Detection Fault', class No Acknowledgement, trigger "DB302_HMI_Faults_Carrier75_Faults_1" bit 0
   4818: 'Carrier 75 Carrier Number Invalid', class No Acknowledgement, trigger "DB302_HMI_Faults_Carrier75_Faults_1" bit 1
   4819: 'Carrier 75 Drive: PROFINET configuration error', class No Acknowledgement, trigger "DB302_HMI_Faults_Carrier75_Faults_1" bit 2
   4820: 'Carrier 75 Drive: Error internal communications', class No Acknowledgement, trigger "DB302_HMI_Faults_Carrier75_Faults_1" bit 3
   4821: 'Carrier 75 Drive: Motor overtemperature', class No Acknowledgement, trigger "DB302_HMI_Faults_Carrier75_Faults_1" bit 4
   4822: 'Carrier 75 Drive: Motor overcurrent', class No Acknowledgement, trigger "DB302_HMI_Faults_Carrier75_Faults_1" bit 5
   4823: 'Carrier 75 Drive: Infeed or power unit not ready', class No Acknowledgement, trigger "DB302_HMI_Faults_Carrier75_Faults_1" bit 6
   4824: 'Carrier 75 Drive: Short-circuit/ground fault detected', class No Acknowledgement, trigger "DB302_HMI_Faults_Carrier75_Faults_1" bit 7
   4825: 'Carrier 75 Drive: PROFINET Setpoint timeout', class No Acknowledgement, trigger "DB302_HMI_Faults_Carrier75_Faults_1" bit 8
   4826: 'Carrier 75 Power unit: Overcurrent', class No Acknowledgement, trigger "DB302_HMI_Faults_Carrier75_Faults_1" bit 9
   4827: 'Carrier 75 Power unit: DC link voltage overvoltage', class No Acknowledgement, trigger "DB302_HMI_Faults_Carrier75_Faults_1" bit 10
   4828: 'Carrier 75 Power unit: DC link voltage undervoltage', class No Acknowledgement, trigger "DB302_HMI_Faults_Carrier75_Faults_1" bit 11
   4829: 'Carrier 75 Power unit: Line phase failure in main circuit', class No Acknowledgement, trigger "DB302_HMI_Faults_Carrier75_Faults_1" bit 12
   4830: 'Carrier 75 Power unit: Phase failure motor cable', class No Acknowledgement, trigger "DB302_HMI_Faults_Carrier75_Faults_1" bit 13
   4831: 'Carrier 75 Power unit: Ground fault', class No Acknowledgement, trigger "DB302_HMI_Faults_Carrier75_Faults_1" bit 14
   4832: 'Spare_Fault_4832', class No Acknowledgement, trigger "DB302_HMI_Faults_Carrier75_Faults_1" bit 15
   4833: 'Carrier 75 Motion Off Fault', class No Acknowledgement, trigger "DB302_HMI_Faults_Carrier75_Faults_2" bit 0
   4834: 'Carrier 75 Motion On Fault', class No Acknowledgement, trigger "DB302_HMI_Faults_Carrier75_Faults_2" bit 1
   4835: 'Carrier 75 Spacing Fault', class No Acknowledgement, trigger "DB302_HMI_Faults_Carrier75_Faults_2" bit 2
   4836: 'Carrier 75 Duplicate Carrier Number Fault', class No Acknowledgement, trigger "DB302_HMI_Faults_Carrier75_Faults_2" bit 3
   4837: 'Spare_Fault_4837', class No Acknowledgement, trigger "DB302_HMI_Faults_Carrier75_Faults_2" bit 4
   4838: 'Spare_Fault_4838', class No Acknowledgement, trigger "DB302_HMI_Faults_Carrier75_Faults_2" bit 5
   4839: 'Spare_Fault_4839', class No Acknowledgement, trigger "DB302_HMI_Faults_Carrier75_Faults_2" bit 6
   4840: 'Spare_Fault_4840', class No Acknowledgement, trigger "DB302_HMI_Faults_Carrier75_Faults_2" bit 7
   4841: 'Spare_Fault_4841', class No Acknowledgement, trigger "DB302_HMI_Faults_Carrier75_Faults_2" bit 8
   4842: 'Spare_Fault_4842', class No Acknowledgement, trigger "DB302_HMI_Faults_Carrier75_Faults_2" bit 9
   4843: 'Spare_Fault_4843', class No Acknowledgement, trigger "DB302_HMI_Faults_Carrier75_Faults_2" bit 10
   4844: 'Spare_Fault_4844', class No Acknowledgement, trigger "DB302_HMI_Faults_Carrier75_Faults_2" bit 11
   4845: 'Spare_Fault_4845', class No Acknowledgement, trigger "DB302_HMI_Faults_Carrier75_Faults_2" bit 12
   4846: 'Spare_Fault_4846', class No Acknowledgement, trigger "DB302_HMI_Faults_Carrier75_Faults_2" bit 13
   4847: 'Spare_Fault_4847', class No Acknowledgement, trigger "DB302_HMI_Faults_Carrier75_Faults_2" bit 14
   4848: 'Spare_Fault_4848', class No Acknowledgement, trigger "DB302_HMI_Faults_Carrier75_Faults_2" bit 15
   4849: 'Spare_Fault_4849', class No Acknowledgement, trigger "DB302_HMI_Faults_Carrier75_Faults_3" bit 0
   4850: 'Spare_Fault_4850', class No Acknowledgement, trigger "DB302_HMI_Faults_Carrier75_Faults_3" bit 1
   4851: 'Spare_Fault_4851', class No Acknowledgement, trigger "DB302_HMI_Faults_Carrier75_Faults_3" bit 2
   4852: 'Spare_Fault_4852', class No Acknowledgement, trigger "DB302_HMI_Faults_Carrier75_Faults_3" bit 3
   4853: 'Spare_Fault_4853', class No Acknowledgement, trigger "DB302_HMI_Faults_Carrier75_Faults_3" bit 4
   4854: 'Spare_Fault_4854', class No Acknowledgement, trigger "DB302_HMI_Faults_Carrier75_Faults_3" bit 5
   4855: 'Spare_Fault_4855', class No Acknowledgement, trigger "DB302_HMI_Faults_Carrier75_Faults_3" bit 6
   4856: 'Spare_Fault_4856', class No Acknowledgement, trigger "DB302_HMI_Faults_Carrier75_Faults_3" bit 7
   4857: 'Spare_Fault_4857', class No Acknowledgement, trigger "DB302_HMI_Faults_Carrier75_Faults_3" bit 8
   4858: 'Spare_Fault_4858', class No Acknowledgement, trigger "DB302_HMI_Faults_Carrier75_Faults_3" bit 9
   4859: 'Spare_Fault_4859', class No Acknowledgement, trigger "DB302_HMI_Faults_Carrier75_Faults_3" bit 10
   4860: 'Spare_Fault_4860', class No Acknowledgement, trigger "DB302_HMI_Faults_Carrier75_Faults_3" bit 11
   4861: 'Spare_Fault_4861', class No Acknowledgement, trigger "DB302_HMI_Faults_Carrier75_Faults_3" bit 12
   4862: 'Spare_Fault_4862', class No Acknowledgement, trigger "DB302_HMI_Faults_Carrier75_Faults_3" bit 13
   4863: 'Spare_Fault_4863', class No Acknowledgement, trigger "DB302_HMI_Faults_Carrier75_Faults_3" bit 14
   4864: 'Spare_Fault_4864', class No Acknowledgement, trigger "DB302_HMI_Faults_Carrier75_Faults_3" bit 15
   4865: 'Carrier 76 Disconnect Open Power Fault DI11.0', class No Acknowledgement, trigger "DB302_HMI_Faults_Carrier76_Faults_0" bit 0
   4866: 'Carrier 76 Drive Profinet Comm Fault', class No Acknowledgement, trigger "DB302_HMI_Faults_Carrier76_Faults_0" bit 1
   4867: 'Carrier 76 Production Stop Not Reset', class No Acknowledgement, trigger "DB302_HMI_Faults_Carrier76_Faults_0" bit 2
   4868: 'Carrier 76 CB02122 Tripped', class No Acknowledgement, trigger "DB302_HMI_Faults_Carrier76_Faults_0" bit 3
   4869: 'Carrier 76 CB02123 Tripped', class No Acknowledgement, trigger "DB302_HMI_Faults_Carrier76_Faults_0" bit 4
   4870: 'Carrier 76 AUX1 CB Tripped', class No Acknowledgement, trigger "DB302_HMI_Faults_Carrier76_Faults_0" bit 5
   4871: 'Carrier 76 AUX2 CB Tripped', class No Acknowledgement, trigger "DB302_HMI_Faults_Carrier76_Faults_0" bit 6
   4872: 'Carrier 76 PLC Not Communicating', class No Acknowledgement, trigger "DB302_HMI_Faults_Carrier76_Faults_0" bit 7
   4873: 'Carrier 76 Safe Input Card Fault', class No Acknowledgement, trigger "DB302_HMI_Faults_Carrier76_Faults_0" bit 8
   4874: 'Carrier 76 Safe Output Card Fault', class No Acknowledgement, trigger "DB302_HMI_Faults_Carrier76_Faults_0" bit 9
   4875: 'Carrier 76 Standard Input Card Fault', class No Acknowledgement, trigger "DB302_HMI_Faults_Carrier76_Faults_0" bit 10
   4876: 'Carrier 76 Standard Output Card Fault', class No Acknowledgement, trigger "DB302_HMI_Faults_Carrier76_Faults_0" bit 11
   4877: 'Carrier 76 Encoder Position Fault', class No Acknowledgement, trigger "DB302_HMI_Faults_Carrier76_Faults_0" bit 12
   4878: 'Carrier 76 Encoder Internal Error', class No Acknowledgement, trigger "DB302_HMI_Faults_Carrier76_Faults_0" bit 13
   4879: 'Carrier 76 Encoder Comm Fault', class No Acknowledgement, trigger "DB302_HMI_Faults_Carrier76_Faults_0" bit 14
   4880: 'Carrier 76 HMI Comm Fault', class No Acknowledgement, trigger "DB302_HMI_Faults_Carrier76_Faults_0" bit 15
   4881: 'Carrier 76 Crash Detection Fault', class No Acknowledgement, trigger "DB302_HMI_Faults_Carrier76_Faults_1" bit 0
   4882: 'Carrier 76 Carrier Number Invalid', class No Acknowledgement, trigger "DB302_HMI_Faults_Carrier76_Faults_1" bit 1
   4883: 'Carrier 76 Drive: PROFINET configuration error', class No Acknowledgement, trigger "DB302_HMI_Faults_Carrier76_Faults_1" bit 2
   4884: 'Carrier 76 Drive: Error internal communications', class No Acknowledgement, trigger "DB302_HMI_Faults_Carrier76_Faults_1" bit 3
   4885: 'Carrier 76 Drive: Motor overtemperature', class No Acknowledgement, trigger "DB302_HMI_Faults_Carrier76_Faults_1" bit 4
   4886: 'Carrier 76 Drive: Motor overcurrent', class No Acknowledgement, trigger "DB302_HMI_Faults_Carrier76_Faults_1" bit 5
   4887: 'Carrier 76 Drive: Infeed or power unit not ready', class No Acknowledgement, trigger "DB302_HMI_Faults_Carrier76_Faults_1" bit 6
   4888: 'Carrier 76 Drive: Short-circuit/ground fault detected', class No Acknowledgement, trigger "DB302_HMI_Faults_Carrier76_Faults_1" bit 7
   4889: 'Carrier 76 Drive: PROFINET Setpoint timeout', class No Acknowledgement, trigger "DB302_HMI_Faults_Carrier76_Faults_1" bit 8
   4890: 'Carrier 76 Power unit: Overcurrent', class No Acknowledgement, trigger "DB302_HMI_Faults_Carrier76_Faults_1" bit 9
   4891: 'Carrier 76 Power unit: DC link voltage overvoltage', class No Acknowledgement, trigger "DB302_HMI_Faults_Carrier76_Faults_1" bit 10
   4892: 'Carrier 76 Power unit: DC link voltage undervoltage', class No Acknowledgement, trigger "DB302_HMI_Faults_Carrier76_Faults_1" bit 11
   4893: 'Carrier 76 Power unit: Line phase failure in main circuit', class No Acknowledgement, trigger "DB302_HMI_Faults_Carrier76_Faults_1" bit 12
   4894: 'Carrier 76 Power unit: Phase failure motor cable', class No Acknowledgement, trigger "DB302_HMI_Faults_Carrier76_Faults_1" bit 13
   4895: 'Carrier 76 Power unit: Ground fault', class No Acknowledgement, trigger "DB302_HMI_Faults_Carrier76_Faults_1" bit 14
   4896: 'Spare_Fault_4896', class No Acknowledgement, trigger "DB302_HMI_Faults_Carrier76_Faults_1" bit 15
   4897: 'Carrier 76 Motion Off Fault', class No Acknowledgement, trigger "DB302_HMI_Faults_Carrier76_Faults_2" bit 0
   4898: 'Carrier 76 Motion On Fault', class No Acknowledgement, trigger "DB302_HMI_Faults_Carrier76_Faults_2" bit 1
   4899: 'Carrier 76 Spacing Fault', class No Acknowledgement, trigger "DB302_HMI_Faults_Carrier76_Faults_2" bit 2
   4900: 'Carrier 76 Duplicate Carrier Number Fault', class No Acknowledgement, trigger "DB302_HMI_Faults_Carrier76_Faults_2" bit 3
   4901: 'Spare_Fault_4901', class No Acknowledgement, trigger "DB302_HMI_Faults_Carrier76_Faults_2" bit 4
   4902: 'Spare_Fault_4902', class No Acknowledgement, trigger "DB302_HMI_Faults_Carrier76_Faults_2" bit 5
   4903: 'Spare_Fault_4903', class No Acknowledgement, trigger "DB302_HMI_Faults_Carrier76_Faults_2" bit 6
   4904: 'Spare_Fault_4904', class No Acknowledgement, trigger "DB302_HMI_Faults_Carrier76_Faults_2" bit 7
   4905: 'Spare_Fault_4905', class No Acknowledgement, trigger "DB302_HMI_Faults_Carrier76_Faults_2" bit 8
   4906: 'Spare_Fault_4906', class No Acknowledgement, trigger "DB302_HMI_Faults_Carrier76_Faults_2" bit 9
   4907: 'Spare_Fault_4907', class No Acknowledgement, trigger "DB302_HMI_Faults_Carrier76_Faults_2" bit 10
   4908: 'Spare_Fault_4908', class No Acknowledgement, trigger "DB302_HMI_Faults_Carrier76_Faults_2" bit 11
   4909: 'Spare_Fault_4909', class No Acknowledgement, trigger "DB302_HMI_Faults_Carrier76_Faults_2" bit 12
